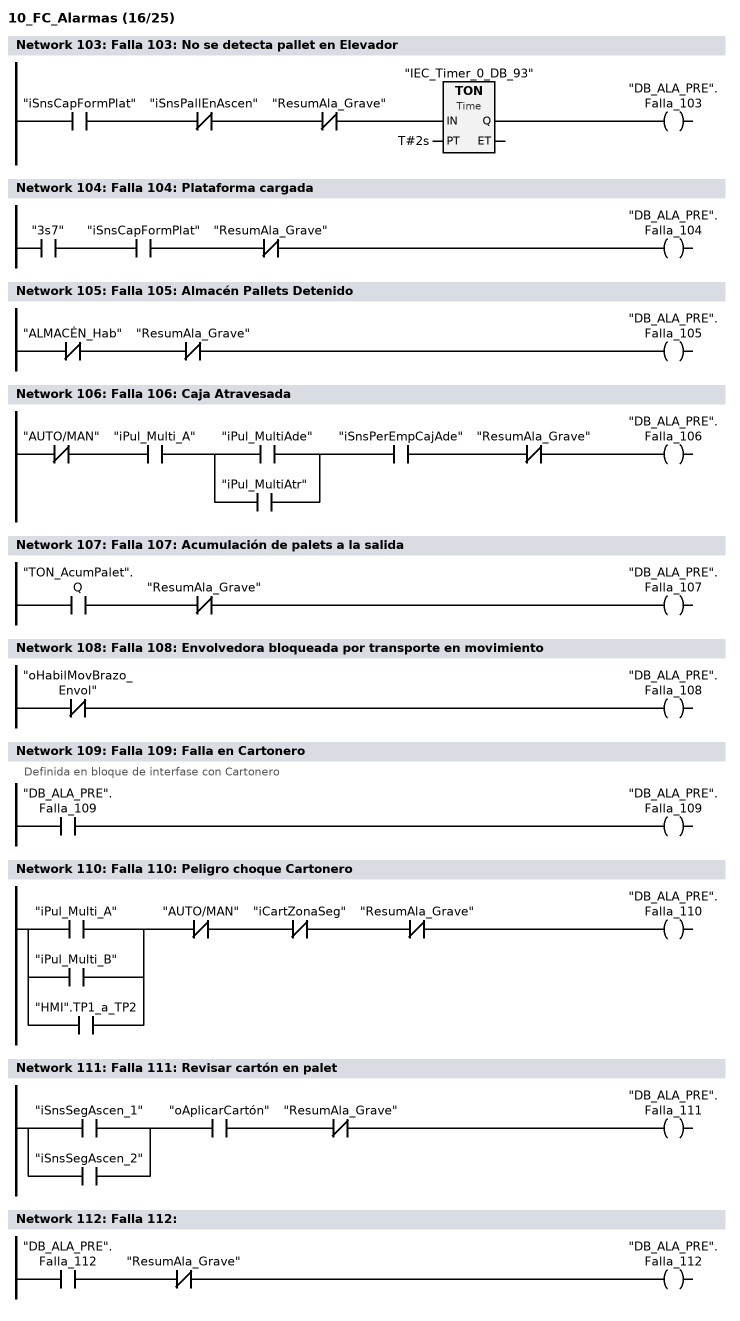
   "IEC_Timer_0_DB_93".TON(IN := "iSnsCapFormPlat" AND NOT "iSnsPallEnAscen" AND NOT "ResumAla_Grave",
                           PT := T#2s);
   "DB_ALA_PRE".Falla_103 := "IEC_Timer_0_DB_93".Q;
END_REGION

REGION Network 104: Falla 104: Plataforma cargada
   RUNG wire#powerrail
      Contact( "3s7" )
      Contact( "iSnsCapFormPlat" )
      I_Contact( "ResumAla_Grave" )
      Coil( "DB_ALA_PRE".Falla_104 )
   END_RUNG
   // the same network as SCL:
   "DB_ALA_PRE".Falla_104 := "3s7" AND "iSnsCapFormPlat" AND NOT "ResumAla_Grave";
END_REGION

REGION Network 105: Falla 105: Almacén Pallets Detenido
   RUNG wire#powerrail
      I_Contact( "ALMACÉN_Hab" )
      I_Contact( "ResumAla_Grave" )
      Coil( "DB_ALA_PRE".Falla_105 )
   END_RUNG
   // the same network as SCL:
   "DB_ALA_PRE".Falla_105 := NOT "ALMACÉN_Hab" AND NOT "ResumAla_Grave";
END_REGION

REGION Network 106: Falla 106: Caja Atravesada
   RUNG wire#powerrail
      I_Contact( "AUTO/MAN" )
      Contact( "iPul_Multi_A" )
      wire#w1
      Contact( "iPul_MultiAde" )
      wire#w2
      Contact( "iSnsPerEmpCajAde" )
      I_Contact( "ResumAla_Grave" )
      Coil( "DB_ALA_PRE".Falla_106 )
   END_RUNG
   RUNG wire#w1
      Contact( "iPul_MultiAtr" )
   END_RUNG wire#w2
   // the same network as SCL:
   "DB_ALA_PRE".Falla_106 := NOT "AUTO/MAN" AND "iPul_Multi_A" AND ("iPul_MultiAde" OR "iPul_MultiAtr") AND "iSnsPerEmpCajAde" AND NOT "ResumAla_Grave";
END_REGION

REGION Network 107: Falla 107: Acumulación de palets a la salida
   RUNG wire#powerrail
      Contact( "TON_AcumPalet".Q )
      I_Contact( "ResumAla_Grave" )
      Coil( "DB_ALA_PRE".Falla_107 )
   END_RUNG
   // the same network as SCL:
   "DB_ALA_PRE".Falla_107 := "TON_AcumPalet".Q AND NOT "ResumAla_Grave";
END_REGION

REGION Network 108: Falla 108: Envolvedora bloqueada por transporte en movimiento
   RUNG wire#powerrail
      I_Contact( "oHabilMovBrazo_Envol" )
      Coil( "DB_ALA_PRE".Falla_108 )
   END_RUNG
   // the same network as SCL:
   "DB_ALA_PRE".Falla_108 := NOT "oHabilMovBrazo_Envol";
END_REGION

REGION Network 109: Falla 109: Falla en Cartonero
   // Definida en bloque de interfase con Cartonero
   RUNG wire#powerrail
      Contact( "DB_ALA_PRE".Falla_109 )
      Coil( "DB_ALA_PRE".Falla_109 )
   END_RUNG
   // the same network as SCL:
   "DB_ALA_PRE".Falla_109 := "DB_ALA_PRE".Falla_109;
END_REGION

REGION Network 110: Falla 110: Peligro choque Cartonero
   RUNG wire#powerrail
      Contact( "iPul_Multi_A" )
      wire#w1
      I_Contact( "AUTO/MAN" )
      I_Contact( "iCartZonaSeg" )
      I_Contact( "ResumAla_Grave" )
      Coil( "DB_ALA_PRE".Falla_110 )
   END_RUNG
   RUNG wire#powerrail
      Contact( "iPul_Multi_B" )
   END_RUNG wire#w1
   RUNG wire#powerrail
      Contact( "HMI".TP1_a_TP2 )
   END_RUNG wire#w1
   // the same network as SCL:
   "DB_ALA_PRE".Falla_110 := ("iPul_Multi_A" OR "iPul_Multi_B" OR "HMI".TP1_a_TP2) AND NOT "AUTO/MAN" AND NOT "iCartZonaSeg" AND NOT "ResumAla_Grave";
END_REGION

REGION Network 111: Falla 111: Revisar cartón en palet
   RUNG wire#powerrail
      Contact( "iSnsSegAscen_1" )
      wire#w1
      Contact( "oAplicarCartón" )
      I_Contact( "ResumAla_Grave" )
      Coil( "DB_ALA_PRE".Falla_111 )
   END_RUNG
   RUNG wire#powerrail
      Contact( "iSnsSegAscen_2" )
   END_RUNG wire#w1
   // the same network as SCL:
   "DB_ALA_PRE".Falla_111 := ("iSnsSegAscen_1" OR "iSnsSegAscen_2") AND "oAplicarCartón" AND NOT "ResumAla_Grave";
END_REGION

REGION Network 112: Falla 112:
   RUNG wire#powerrail
      Contact( "DB_ALA_PRE".Falla_112 )
      I_Contact( "ResumAla_Grave" )
      Coil( "DB_ALA_PRE".Falla_112 )
   END_RUNG
   // the same network as SCL:
   "DB_ALA_PRE".Falla_112 := "DB_ALA_PRE".Falla_112 AND NOT "ResumAla_Grave";
END_REGION

REGION Network 113: Falla 113: Falla confirm. K18: Empujador Filas Subir
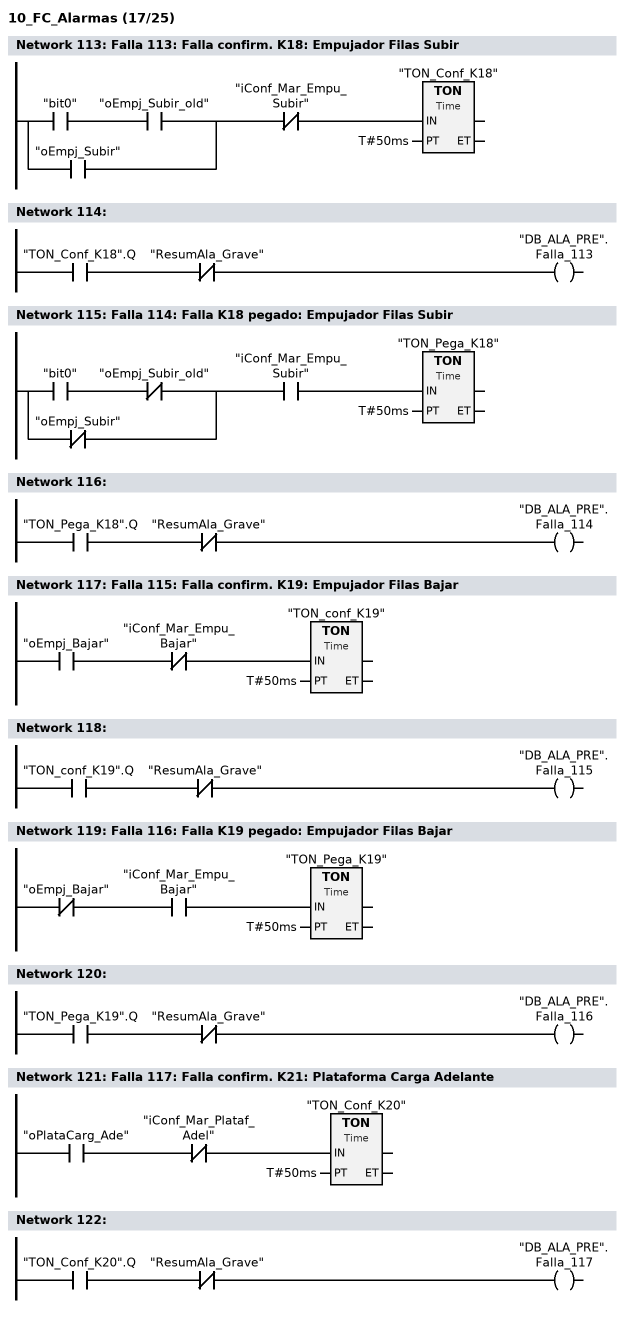
   "TON_Conf_K18".TON(IN := (("bit0" AND "oEmpj_Subir_old") OR "oEmpj_Subir") AND NOT "iConf_Mar_Empu_Subir",
                      PT := T#50ms);
END_REGION

REGION Network 114
   RUNG wire#powerrail
      Contact( "TON_Conf_K18".Q )
      I_Contact( "ResumAla_Grave" )
      Coil( "DB_ALA_PRE".Falla_113 )
   END_RUNG
   // the same network as SCL:
   "DB_ALA_PRE".Falla_113 := "TON_Conf_K18".Q AND NOT "ResumAla_Grave";
END_REGION

REGION Network 115: Falla 114: Falla K18 pegado: Empujador Filas Subir
   "TON_Pega_K18".TON(IN := (("bit0" AND NOT "oEmpj_Subir_old") OR NOT "oEmpj_Subir") AND "iConf_Mar_Empu_Subir",
                      PT := T#50ms);
END_REGION

REGION Network 116
   RUNG wire#powerrail
      Contact( "TON_Pega_K18".Q )
      I_Contact( "ResumAla_Grave" )
      Coil( "DB_ALA_PRE".Falla_114 )
   END_RUNG
   // the same network as SCL:
   "DB_ALA_PRE".Falla_114 := "TON_Pega_K18".Q AND NOT "ResumAla_Grave";
END_REGION

REGION Network 117: Falla 115: Falla confirm. K19: Empujador Filas Bajar
   "TON_conf_K19".TON(IN := "oEmpj_Bajar" AND NOT "iConf_Mar_Empu_Bajar", PT := T#50ms);
END_REGION

REGION Network 118
   RUNG wire#powerrail
      Contact( "TON_conf_K19".Q )
      I_Contact( "ResumAla_Grave" )
      Coil( "DB_ALA_PRE".Falla_115 )
   END_RUNG
   // the same network as SCL:
   "DB_ALA_PRE".Falla_115 := "TON_conf_K19".Q AND NOT "ResumAla_Grave";
END_REGION

REGION Network 119: Falla 116: Falla K19 pegado: Empujador Filas Bajar
   "TON_Pega_K19".TON(IN := NOT "oEmpj_Bajar" AND "iConf_Mar_Empu_Bajar", PT := T#50ms);
END_REGION

REGION Network 120
   RUNG wire#powerrail
      Contact( "TON_Pega_K19".Q )
      I_Contact( "ResumAla_Grave" )
      Coil( "DB_ALA_PRE".Falla_116 )
   END_RUNG
   // the same network as SCL:
   "DB_ALA_PRE".Falla_116 := "TON_Pega_K19".Q AND NOT "ResumAla_Grave";
END_REGION

REGION Network 121: Falla 117: Falla confirm. K21: Plataforma Carga Adelante
   "TON_Conf_K20".TON(IN := "oPlataCarg_Ade" AND NOT "iConf_Mar_Plataf_Adel", PT := T#50ms);
END_REGION

REGION Network 122
   RUNG wire#powerrail
      Contact( "TON_Conf_K20".Q )
      I_Contact( "ResumAla_Grave" )
      Coil( "DB_ALA_PRE".Falla_117 )
   END_RUNG
   // the same network as SCL:
   "DB_ALA_PRE".Falla_117 := "TON_Conf_K20".Q AND NOT "ResumAla_Grave";
END_REGION

REGION Network 123: Falla 118: Falla K21 pegado: Plataforma Carga Adelante
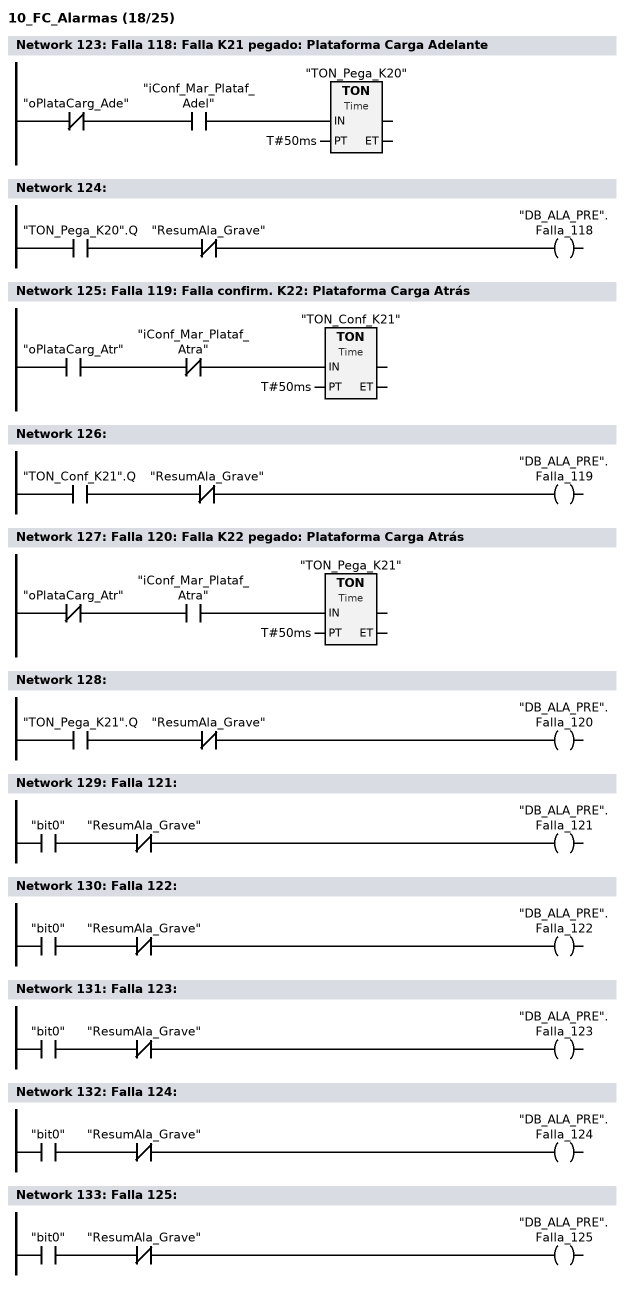
   "TON_Pega_K20".TON(IN := NOT "oPlataCarg_Ade" AND "iConf_Mar_Plataf_Adel", PT := T#50ms);
END_REGION

REGION Network 124
   RUNG wire#powerrail
      Contact( "TON_Pega_K20".Q )
      I_Contact( "ResumAla_Grave" )
      Coil( "DB_ALA_PRE".Falla_118 )
   END_RUNG
   // the same network as SCL:
   "DB_ALA_PRE".Falla_118 := "TON_Pega_K20".Q AND NOT "ResumAla_Grave";
END_REGION

REGION Network 125: Falla 119: Falla confirm. K22: Plataforma Carga Atrás
   "TON_Conf_K21".TON(IN := "oPlataCarg_Atr" AND NOT "iConf_Mar_Plataf_Atra", PT := T#50ms);
END_REGION

REGION Network 126
   RUNG wire#powerrail
      Contact( "TON_Conf_K21".Q )
      I_Contact( "ResumAla_Grave" )
      Coil( "DB_ALA_PRE".Falla_119 )
   END_RUNG
   // the same network as SCL:
   "DB_ALA_PRE".Falla_119 := "TON_Conf_K21".Q AND NOT "ResumAla_Grave";
END_REGION

REGION Network 127: Falla 120: Falla K22 pegado: Plataforma Carga Atrás
   "TON_Pega_K21".TON(IN := NOT "oPlataCarg_Atr" AND "iConf_Mar_Plataf_Atra", PT := T#50ms);
END_REGION

REGION Network 128
   RUNG wire#powerrail
      Contact( "TON_Pega_K21".Q )
      I_Contact( "ResumAla_Grave" )
      Coil( "DB_ALA_PRE".Falla_120 )
   END_RUNG
   // the same network as SCL:
   "DB_ALA_PRE".Falla_120 := "TON_Pega_K21".Q AND NOT "ResumAla_Grave";
END_REGION

REGION Network 129: Falla 121:
   RUNG wire#powerrail
      Contact( "bit0" )
      I_Contact( "ResumAla_Grave" )
      Coil( "DB_ALA_PRE".Falla_121 )
   END_RUNG
   // the same network as SCL:
   "DB_ALA_PRE".Falla_121 := "bit0" AND NOT "ResumAla_Grave";
END_REGION

REGION Network 130: Falla 122:
   RUNG wire#powerrail
      Contact( "bit0" )
      I_Contact( "ResumAla_Grave" )
      Coil( "DB_ALA_PRE".Falla_122 )
   END_RUNG
   // the same network as SCL:
   "DB_ALA_PRE".Falla_122 := "bit0" AND NOT "ResumAla_Grave";
END_REGION

REGION Network 131: Falla 123:
   RUNG wire#powerrail
      Contact( "bit0" )
      I_Contact( "ResumAla_Grave" )
      Coil( "DB_ALA_PRE".Falla_123 )
   END_RUNG
   // the same network as SCL:
   "DB_ALA_PRE".Falla_123 := "bit0" AND NOT "ResumAla_Grave";
END_REGION

REGION Network 132: Falla 124:
   RUNG wire#powerrail
      Contact( "bit0" )
      I_Contact( "ResumAla_Grave" )
      Coil( "DB_ALA_PRE".Falla_124 )
   END_RUNG
   // the same network as SCL:
   "DB_ALA_PRE".Falla_124 := "bit0" AND NOT "ResumAla_Grave";
END_REGION

REGION Network 133: Falla 125:
   RUNG wire#powerrail
      Contact( "bit0" )
      I_Contact( "ResumAla_Grave" )
      Coil( "DB_ALA_PRE".Falla_125 )
   END_RUNG
   // the same network as SCL:
   "DB_ALA_PRE".Falla_125 := "bit0" AND NOT "ResumAla_Grave";
END_REGION

REGION Network 134: Falla 126:
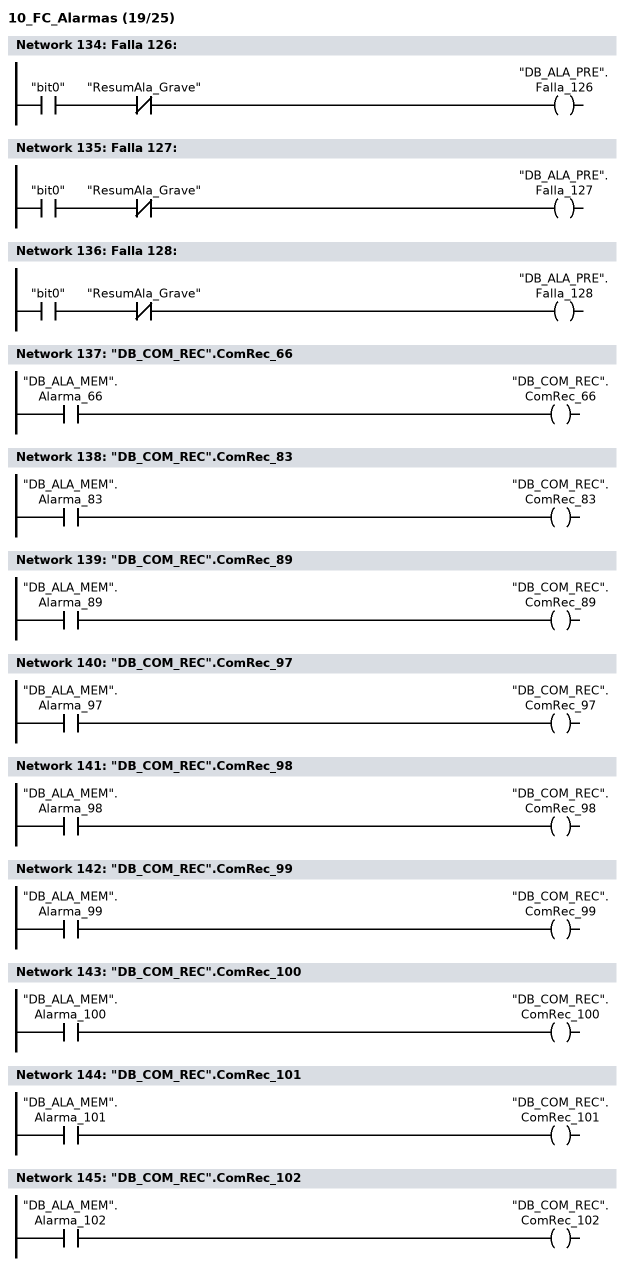
   RUNG wire#powerrail
      Contact( "bit0" )
      I_Contact( "ResumAla_Grave" )
      Coil( "DB_ALA_PRE".Falla_126 )
   END_RUNG
   // the same network as SCL:
   "DB_ALA_PRE".Falla_126 := "bit0" AND NOT "ResumAla_Grave";
END_REGION

REGION Network 135: Falla 127:
   RUNG wire#powerrail
      Contact( "bit0" )
      I_Contact( "ResumAla_Grave" )
      Coil( "DB_ALA_PRE".Falla_127 )
   END_RUNG
   // the same network as SCL:
   "DB_ALA_PRE".Falla_127 := "bit0" AND NOT "ResumAla_Grave";
END_REGION

REGION Network 136: Falla 128:
   RUNG wire#powerrail
      Contact( "bit0" )
      I_Contact( "ResumAla_Grave" )
      Coil( "DB_ALA_PRE".Falla_128 )
   END_RUNG
   // the same network as SCL:
   "DB_ALA_PRE".Falla_128 := "bit0" AND NOT "ResumAla_Grave";
END_REGION

REGION Network 137: "DB_COM_REC".ComRec_66
   RUNG wire#powerrail
      Contact( "DB_ALA_MEM".Alarma_66 )
      Coil( "DB_COM_REC".ComRec_66 )
   END_RUNG
   // the same network as SCL:
   "DB_COM_REC".ComRec_66 := "DB_ALA_MEM".Alarma_66;
END_REGION

REGION Network 138: "DB_COM_REC".ComRec_83
   RUNG wire#powerrail
      Contact( "DB_ALA_MEM".Alarma_83 )
      Coil( "DB_COM_REC".ComRec_83 )
   END_RUNG
   // the same network as SCL:
   "DB_COM_REC".ComRec_83 := "DB_ALA_MEM".Alarma_83;
END_REGION

REGION Network 139: "DB_COM_REC".ComRec_89
   RUNG wire#powerrail
      Contact( "DB_ALA_MEM".Alarma_89 )
      Coil( "DB_COM_REC".ComRec_89 )
   END_RUNG
   // the same network as SCL:
   "DB_COM_REC".ComRec_89 := "DB_ALA_MEM".Alarma_89;
END_REGION

REGION Network 140: "DB_COM_REC".ComRec_97
   RUNG wire#powerrail
      Contact( "DB_ALA_MEM".Alarma_97 )
      Coil( "DB_COM_REC".ComRec_97 )
   END_RUNG
   // the same network as SCL:
   "DB_COM_REC".ComRec_97 := "DB_ALA_MEM".Alarma_97;
END_REGION

REGION Network 141: "DB_COM_REC".ComRec_98
   RUNG wire#powerrail
      Contact( "DB_ALA_MEM".Alarma_98 )
      Coil( "DB_COM_REC".ComRec_98 )
   END_RUNG
   // the same network as SCL:
   "DB_COM_REC".ComRec_98 := "DB_ALA_MEM".Alarma_98;
END_REGION

REGION Network 142: "DB_COM_REC".ComRec_99
   RUNG wire#powerrail
      Contact( "DB_ALA_MEM".Alarma_99 )
      Coil( "DB_COM_REC".ComRec_99 )
   END_RUNG
   // the same network as SCL:
   "DB_COM_REC".ComRec_99 := "DB_ALA_MEM".Alarma_99;
END_REGION

REGION Network 143: "DB_COM_REC".ComRec_100
   RUNG wire#powerrail
      Contact( "DB_ALA_MEM".Alarma_100 )
      Coil( "DB_COM_REC".ComRec_100 )
   END_RUNG
   // the same network as SCL:
   "DB_COM_REC".ComRec_100 := "DB_ALA_MEM".Alarma_100;
END_REGION

REGION Network 144: "DB_COM_REC".ComRec_101
   RUNG wire#powerrail
      Contact( "DB_ALA_MEM".Alarma_101 )
      Coil( "DB_COM_REC".ComRec_101 )
   END_RUNG
   // the same network as SCL:
   "DB_COM_REC".ComRec_101 := "DB_ALA_MEM".Alarma_101;
END_REGION

REGION Network 145: "DB_COM_REC".ComRec_102
   RUNG wire#powerrail
      Contact( "DB_ALA_MEM".Alarma_102 )
      Coil( "DB_COM_REC".ComRec_102 )
   END_RUNG
   // the same network as SCL:
   "DB_COM_REC".ComRec_102 := "DB_ALA_MEM".Alarma_102;
END_REGION

REGION Network 146: "DB_COM_REC".ComRec_103
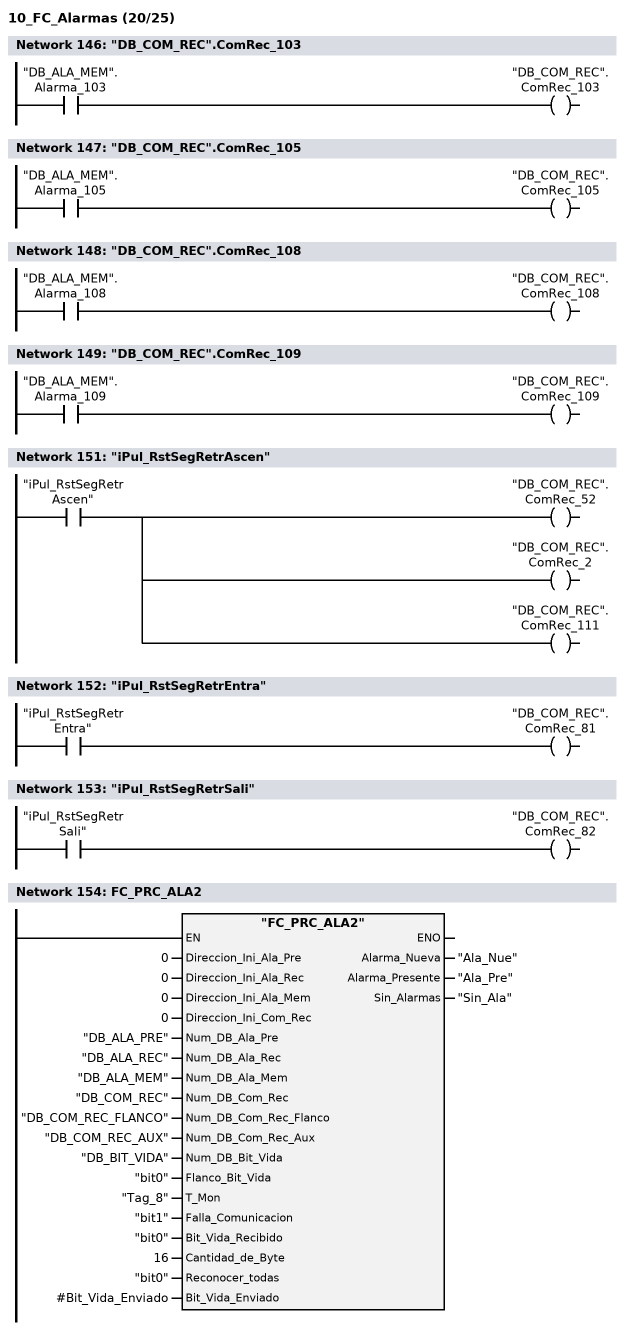
   RUNG wire#powerrail
      Contact( "DB_ALA_MEM".Alarma_103 )
      Coil( "DB_COM_REC".ComRec_103 )
   END_RUNG
   // the same network as SCL:
   "DB_COM_REC".ComRec_103 := "DB_ALA_MEM".Alarma_103;
END_REGION

REGION Network 147: "DB_COM_REC".ComRec_105
   RUNG wire#powerrail
      Contact( "DB_ALA_MEM".Alarma_105 )
      Coil( "DB_COM_REC".ComRec_105 )
   END_RUNG
   // the same network as SCL:
   "DB_COM_REC".ComRec_105 := "DB_ALA_MEM".Alarma_105;
END_REGION

REGION Network 148: "DB_COM_REC".ComRec_108
   RUNG wire#powerrail
      Contact( "DB_ALA_MEM".Alarma_108 )
      Coil( "DB_COM_REC".ComRec_108 )
   END_RUNG
   // the same network as SCL:
   "DB_COM_REC".ComRec_108 := "DB_ALA_MEM".Alarma_108;
END_REGION

REGION Network 149: "DB_COM_REC".ComRec_109
   RUNG wire#powerrail
      Contact( "DB_ALA_MEM".Alarma_109 )
      Coil( "DB_COM_REC".ComRec_109 )
   END_RUNG
   // the same network as SCL:
   "DB_COM_REC".ComRec_109 := "DB_ALA_MEM".Alarma_109;
END_REGION

REGION Network 150: ------------------------------------------------------------------------------------------------------------------------------------------------------------------------------------------------------
END_REGION

REGION Network 151: "iPul_RstSegRetrAscen"
   RUNG wire#powerrail
      Contact( "iPul_RstSegRetrAscen" )
      wire#w1
      Coil( "DB_COM_REC".ComRec_52 )
   END_RUNG
   RUNG wire#w1
      Coil( "DB_COM_REC".ComRec_2 )
   END_RUNG
   RUNG wire#w1
      Coil( "DB_COM_REC".ComRec_111 )
   END_RUNG
   // the same network as SCL:
   "DB_COM_REC".ComRec_52 := "iPul_RstSegRetrAscen";
   "DB_COM_REC".ComRec_2 := "iPul_RstSegRetrAscen";
   "DB_COM_REC".ComRec_111 := "iPul_RstSegRetrAscen";
END_REGION

REGION Network 152: "iPul_RstSegRetrEntra"
   RUNG wire#powerrail
      Contact( "iPul_RstSegRetrEntra" )
      Coil( "DB_COM_REC".ComRec_81 )
   END_RUNG
   // the same network as SCL:
   "DB_COM_REC".ComRec_81 := "iPul_RstSegRetrEntra";
END_REGION

REGION Network 153: "iPul_RstSegRetrSali"
   RUNG wire#powerrail
      Contact( "iPul_RstSegRetrSali" )
      Coil( "DB_COM_REC".ComRec_82 )
   END_RUNG
   // the same network as SCL:
   "DB_COM_REC".ComRec_82 := "iPul_RstSegRetrSali";
END_REGION

REGION Network 154: FC_PRC_ALA2
   RUNG wire#powerrail
      "FC_PRC_ALA2"(Direccion_Ini_Ala_Pre := 0, Direccion_Ini_Ala_Rec := 0, Direccion_Ini_Ala_Mem := 0, Direccion_Ini_Com_Rec := 0, Num_DB_Ala_Pre := "DB_ALA_PRE", Num_DB_Ala_Rec := "DB_ALA_REC", Num_DB_Ala_Mem := "DB_ALA_MEM", Num_DB_Com_Rec := "DB_COM_REC", Num_DB_Com_Rec_Flanco := "DB_COM_REC_FLANCO", Num_DB_Com_Rec_Aux := "DB_COM_REC_AUX", Num_DB_Bit_Vida := "DB_BIT_VIDA", Flanco_Bit_Vida := "bit0", T_Mon := "Tag_8", Falla_Comunicacion := "bit1", Bit_Vida_Recibido := "bit0", Cantidad_de_Byte := 16, Reconocer_todas := "bit0", Bit_Vida_Enviado := #Bit_Vida_Enviado, Alarma_Nueva => "Ala_Nue", Alarma_Presente => "Ala_Pre", Sin_Alarmas => "Sin_Ala")
   END_RUNG
   // the same network as SCL:
   "FC_PRC_ALA2"(Direccion_Ini_Ala_Pre := 0,
                 Direccion_Ini_Ala_Rec := 0,
                 Direccion_Ini_Ala_Mem := 0,
                 Direccion_Ini_Com_Rec := 0,
                 Num_DB_Ala_Pre := "DB_ALA_PRE",
                 Num_DB_Ala_Rec := "DB_ALA_REC",
                 Num_DB_Ala_Mem := "DB_ALA_MEM",
                 Num_DB_Com_Rec := "DB_COM_REC",
                 Num_DB_Com_Rec_Flanco := "DB_COM_REC_FLANCO",
                 Num_DB_Com_Rec_Aux := "DB_COM_REC_AUX",
                 Num_DB_Bit_Vida := "DB_BIT_VIDA",
                 Flanco_Bit_Vida := "bit0",
                 T_Mon := "Tag_8",
                 Falla_Comunicacion := "bit1",
                 Bit_Vida_Recibido := "bit0",
                 Cantidad_de_Byte := 16,
                 Reconocer_todas := "bit0",
                 Bit_Vida_Enviado := #Bit_Vida_Enviado,
                 Alarma_Nueva => "Ala_Nue",
                 Alarma_Presente => "Ala_Pre",
                 Sin_Alarmas => "Sin_Ala");
END_REGION

REGION Network 155: --------------------------------------------------------------------------------------------------------------------------------------------------------------------------------------------------
END_REGION

REGION Network 156: "ResumAla_Grave"
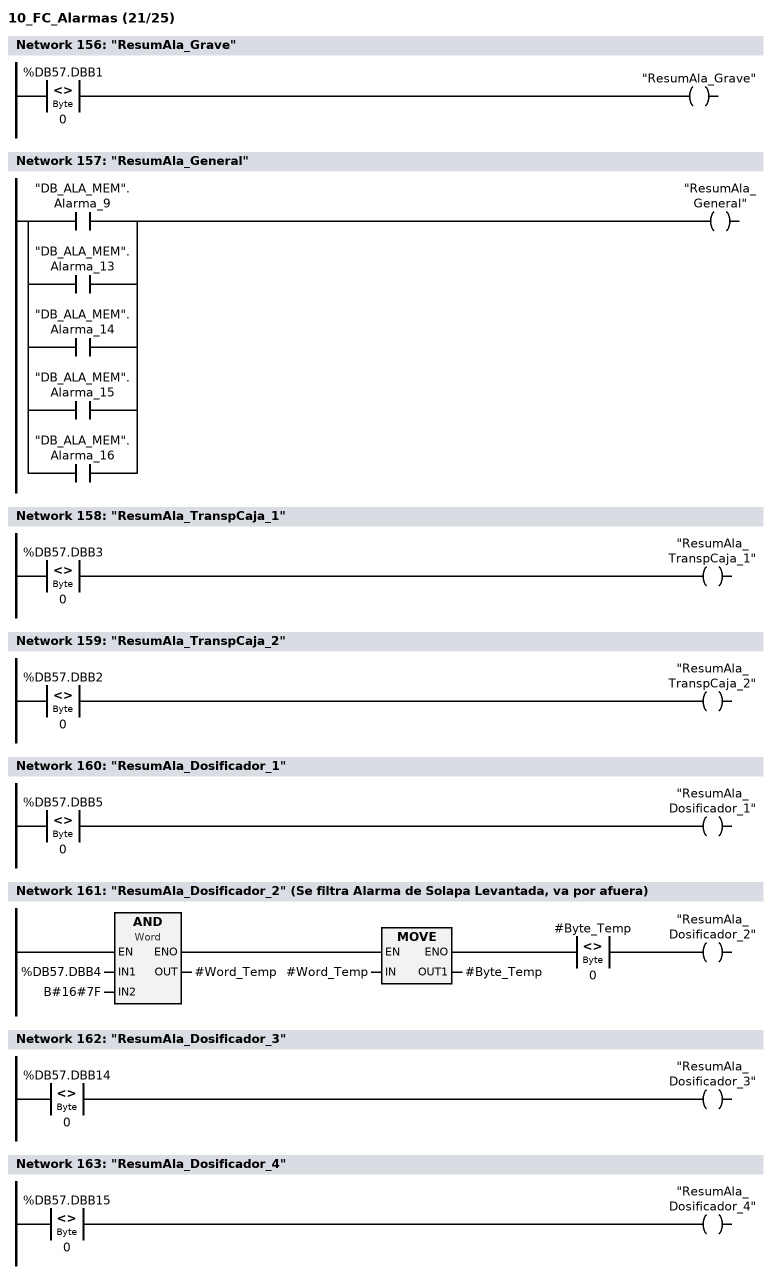
   RUNG wire#powerrail
      { S7_Templates := "SrcType := Byte" } NE_Contact(in1 := %DB57.DBB1, in2 := 0)
      Coil( "ResumAla_Grave" )
   END_RUNG
   // the same network as SCL:
   "ResumAla_Grave" := %DB57.DBB1 <> 0;
END_REGION

REGION Network 157: "ResumAla_General"
   RUNG wire#powerrail
      Contact( "DB_ALA_MEM".Alarma_9 )
      wire#w1
      Coil( "ResumAla_General" )
   END_RUNG
   RUNG wire#powerrail
      Contact( "DB_ALA_MEM".Alarma_13 )
   END_RUNG wire#w1
   RUNG wire#powerrail
      Contact( "DB_ALA_MEM".Alarma_14 )
   END_RUNG wire#w1
   RUNG wire#powerrail
      Contact( "DB_ALA_MEM".Alarma_15 )
   END_RUNG wire#w1
   RUNG wire#powerrail
      Contact( "DB_ALA_MEM".Alarma_16 )
   END_RUNG wire#w1
   // the same network as SCL:
   "ResumAla_General" := "DB_ALA_MEM".Alarma_9 OR "DB_ALA_MEM".Alarma_13 OR "DB_ALA_MEM".Alarma_14 OR "DB_ALA_MEM".Alarma_15 OR "DB_ALA_MEM".Alarma_16;
END_REGION

REGION Network 158: "ResumAla_TranspCaja_1"
   RUNG wire#powerrail
      { S7_Templates := "SrcType := Byte" } NE_Contact(in1 := %DB57.DBB3, in2 := 0)
      Coil( "ResumAla_TranspCaja_1" )
   END_RUNG
   // the same network as SCL:
   "ResumAla_TranspCaja_1" := %DB57.DBB3 <> 0;
END_REGION

REGION Network 159: "ResumAla_TranspCaja_2"
   RUNG wire#powerrail
      { S7_Templates := "SrcType := Byte" } NE_Contact(in1 := %DB57.DBB2, in2 := 0)
      Coil( "ResumAla_TranspCaja_2" )
   END_RUNG
   // the same network as SCL:
   "ResumAla_TranspCaja_2" := %DB57.DBB2 <> 0;
END_REGION

REGION Network 160: "ResumAla_Dosificador_1"
   RUNG wire#powerrail
      { S7_Templates := "SrcType := Byte" } NE_Contact(in1 := %DB57.DBB5, in2 := 0)
      Coil( "ResumAla_Dosificador_1" )
   END_RUNG
   // the same network as SCL:
   "ResumAla_Dosificador_1" := %DB57.DBB5 <> 0;
END_REGION

REGION Network 161: "ResumAla_Dosificador_2" (Se filtra Alarma de Solapa Levantada, va por afuera)
   // no checked SCL form for this network; see the picture
END_REGION

REGION Network 162: "ResumAla_Dosificador_3"
   RUNG wire#powerrail
      { S7_Templates := "SrcType := Byte" } NE_Contact(in1 := %DB57.DBB14, in2 := 0)
      Coil( "ResumAla_Dosificador_3" )
   END_RUNG
   // the same network as SCL:
   "ResumAla_Dosificador_3" := %DB57.DBB14 <> 0;
END_REGION

REGION Network 163: "ResumAla_Dosificador_4"
   RUNG wire#powerrail
      { S7_Templates := "SrcType := Byte" } NE_Contact(in1 := %DB57.DBB15, in2 := 0)
      Coil( "ResumAla_Dosificador_4" )
   END_RUNG
   // the same network as SCL:
   "ResumAla_Dosificador_4" := %DB57.DBB15 <> 0;
END_REGION

REGION Network 164: "ResumAla_CargaPallet_1"
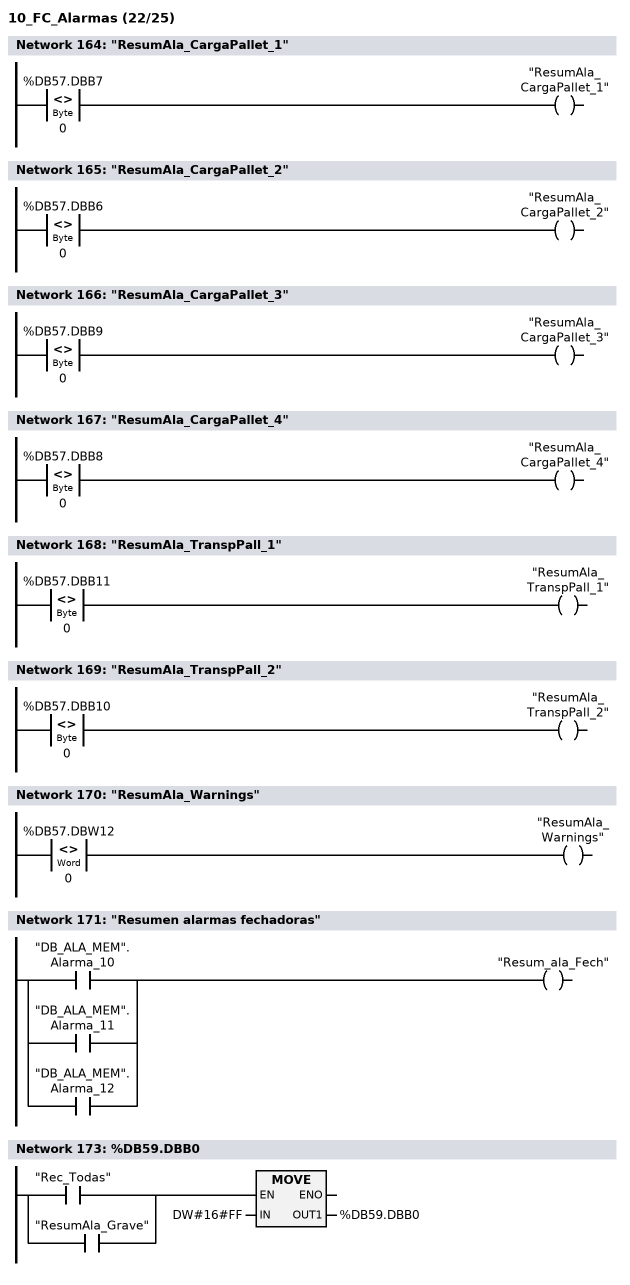
   RUNG wire#powerrail
      { S7_Templates := "SrcType := Byte" } NE_Contact(in1 := %DB57.DBB7, in2 := 0)
      Coil( "ResumAla_CargaPallet_1" )
   END_RUNG
   // the same network as SCL:
   "ResumAla_CargaPallet_1" := %DB57.DBB7 <> 0;
END_REGION

REGION Network 165: "ResumAla_CargaPallet_2"
   RUNG wire#powerrail
      { S7_Templates := "SrcType := Byte" } NE_Contact(in1 := %DB57.DBB6, in2 := 0)
      Coil( "ResumAla_CargaPallet_2" )
   END_RUNG
   // the same network as SCL:
   "ResumAla_CargaPallet_2" := %DB57.DBB6 <> 0;
END_REGION

REGION Network 166: "ResumAla_CargaPallet_3"
   RUNG wire#powerrail
      { S7_Templates := "SrcType := Byte" } NE_Contact(in1 := %DB57.DBB9, in2 := 0)
      Coil( "ResumAla_CargaPallet_3" )
   END_RUNG
   // the same network as SCL:
   "ResumAla_CargaPallet_3" := %DB57.DBB9 <> 0;
END_REGION

REGION Network 167: "ResumAla_CargaPallet_4"
   RUNG wire#powerrail
      { S7_Templates := "SrcType := Byte" } NE_Contact(in1 := %DB57.DBB8, in2 := 0)
      Coil( "ResumAla_CargaPallet_4" )
   END_RUNG
   // the same network as SCL:
   "ResumAla_CargaPallet_4" := %DB57.DBB8 <> 0;
END_REGION

REGION Network 168: "ResumAla_TranspPall_1"
   RUNG wire#powerrail
      { S7_Templates := "SrcType := Byte" } NE_Contact(in1 := %DB57.DBB11, in2 := 0)
      Coil( "ResumAla_TranspPall_1" )
   END_RUNG
   // the same network as SCL:
   "ResumAla_TranspPall_1" := %DB57.DBB11 <> 0;
END_REGION

REGION Network 169: "ResumAla_TranspPall_2"
   RUNG wire#powerrail
      { S7_Templates := "SrcType := Byte" } NE_Contact(in1 := %DB57.DBB10, in2 := 0)
      Coil( "ResumAla_TranspPall_2" )
   END_RUNG
   // the same network as SCL:
   "ResumAla_TranspPall_2" := %DB57.DBB10 <> 0;
END_REGION

REGION Network 170: "ResumAla_Warnings"
   RUNG wire#powerrail
      { S7_Templates := "SrcType := Word" } NE_Contact(in1 := %DB57.DBW12, in2 := 0)
      Coil( "ResumAla_Warnings" )
   END_RUNG
   // the same network as SCL:
   "ResumAla_Warnings" := %DB57.DBW12 <> 0;
END_REGION

REGION Network 171: "Resumen alarmas fechadoras"
   RUNG wire#powerrail
      Contact( "DB_ALA_MEM".Alarma_10 )
      wire#w1
      Coil( "Resum_ala_Fech" )
   END_RUNG
   RUNG wire#powerrail
      Contact( "DB_ALA_MEM".Alarma_11 )
   END_RUNG wire#w1
   RUNG wire#powerrail
      Contact( "DB_ALA_MEM".Alarma_12 )
   END_RUNG wire#w1
   // the same network as SCL:
   "Resum_ala_Fech" := "DB_ALA_MEM".Alarma_10 OR "DB_ALA_MEM".Alarma_11 OR "DB_ALA_MEM".Alarma_12;
END_REGION

REGION Network 172: ------------------------------------------------------------------------------------------------------------------------------------------------------------------------------------------------------
END_REGION

REGION Network 173: %DB59.DBB0
   RUNG wire#powerrail
      Contact( "Rec_Todas" )
      wire#w1
      { S7_GenerateENO := "TRUE" } Move(in := DW#16#FF, out1 => %DB59.DBB0)
   END_RUNG
   RUNG wire#powerrail
      Contact( "ResumAla_Grave" )
   END_RUNG wire#w1
   // the same network as SCL:
   IF "Rec_Todas" OR "ResumAla_Grave" THEN %DB59.DBB0 := DW#16#FF; END_IF;
END_REGION

REGION Network 174: %DB59.DBD0
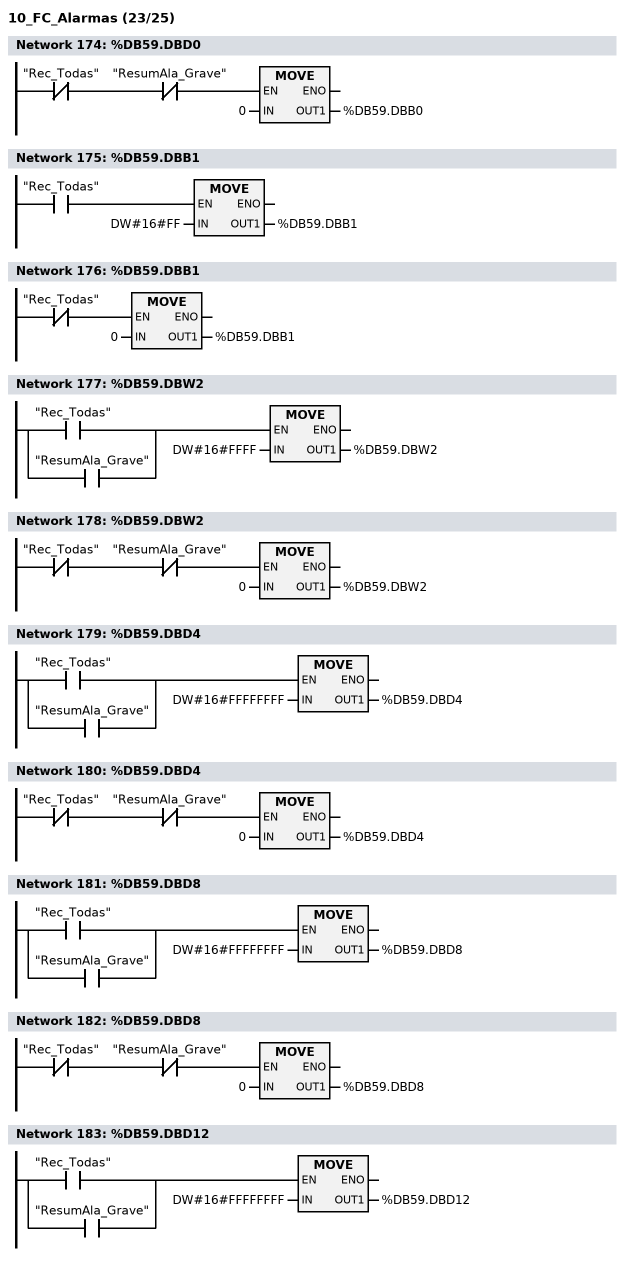
   RUNG wire#powerrail
      I_Contact( "Rec_Todas" )
      I_Contact( "ResumAla_Grave" )
      { S7_GenerateENO := "TRUE" } Move(in := 0, out1 => %DB59.DBB0)
   END_RUNG
   // the same network as SCL:
   IF NOT "Rec_Todas" AND NOT "ResumAla_Grave" THEN %DB59.DBB0 := 0; END_IF;
END_REGION

REGION Network 175: %DB59.DBB1
   RUNG wire#powerrail
      Contact( "Rec_Todas" )
      { S7_GenerateENO := "TRUE" } Move(in := DW#16#FF, out1 => %DB59.DBB1)
   END_RUNG
   // the same network as SCL:
   IF "Rec_Todas" THEN %DB59.DBB1 := DW#16#FF; END_IF;
END_REGION

REGION Network 176: %DB59.DBB1
   RUNG wire#powerrail
      I_Contact( "Rec_Todas" )
      { S7_GenerateENO := "TRUE" } Move(in := 0, out1 => %DB59.DBB1)
   END_RUNG
   // the same network as SCL:
   IF NOT "Rec_Todas" THEN %DB59.DBB1 := 0; END_IF;
END_REGION
